
HMI tags "Consumtion"
   "DB_Zaehler_Anzeige_ViewPreShift" : Bool = PLC DB_Zaehler_Anzeige.ViewPreShift AT %DB211.DBX4.4, 1 s
   "DB_Zaehler_Anzeige_ReadWriteDeviceNo" : Int = PLC DB_Zaehler_Anzeige.ReadWriteDeviceNo AT %DB211.DBW0, 1 s
   "DB_Zaehler_Anzeige_Gesamt_Anzahl" : Int = PLC DB_Zaehler_Anzeige.Gesamt.Anzahl AT %DB211.DBW6, 1 s
   "DB_Zaehler_Anzeige_Gesamt_Verbrauch_K1" : Real = PLC DB_Zaehler_Anzeige.Gesamt.Verbrauch_K1 AT %DB211.DBD8, 1 s
   "DB_Zaehler_Anzeige_Gesamt_Verbrauch_K2" : Real = PLC DB_Zaehler_Anzeige.Gesamt.Verbrauch_K2 AT %DB211.DBD12, 1 s
   "DB_Zaehler_Anzeige_Gesamt_Verbrauch_K3" : Real = PLC DB_Zaehler_Anzeige.Gesamt.Verbrauch_K3 AT %DB211.DBD16, 1 s
   "DB_Zaehler_Anzeige_Gesamt_Verbrauch_K4" : Real = PLC DB_Zaehler_Anzeige.Gesamt.Verbrauch_K4 AT %DB211.DBD20, 1 s
   "DB_Zaehler_Anzeige_Gesamt_Verbrauch_K5" : Real = PLC DB_Zaehler_Anzeige.Gesamt.Verbrauch_K5 AT %DB211.DBD24, 1 s
   "DB_Zaehler_Anzeige_Gesamt_Verbrauch_K6" : Real = PLC DB_Zaehler_Anzeige.Gesamt.Verbrauch_K6 AT %DB211.DBD28, 1 s
   "DB_Zaehler_Anzeige_Gesamt_Verbrauch_K7" : Real = PLC DB_Zaehler_Anzeige.Gesamt.Verbrauch_K7 AT %DB211.DBD32, 1 s
   "DB_Zaehler_Anzeige_Gesamt_Verbrauch_K8" : Real = PLC DB_Zaehler_Anzeige.Gesamt.Verbrauch_K8 AT %DB211.DBD36, 1 s
   "DB_Zaehler_Anzeige_Counter{1}_Anzahl" : Int = PLC DB_Zaehler_Anzeige.Counter[1].Anzahl AT %DB211.DBW40, 1 s
   "DB_Zaehler_Anzeige_Counter{1}_Verbrauch_K1" : Real = PLC DB_Zaehler_Anzeige.Counter[1].Verbrauch_K1 AT %DB211.DBD42, 1 s
   "DB_Zaehler_Anzeige_Counter{1}_Verbrauch_K2" : Real = PLC DB_Zaehler_Anzeige.Counter[1].Verbrauch_K2 AT %DB211.DBD46, 1 s
   "DB_Zaehler_Anzeige_Counter{1}_Verbrauch_K3" : Real = PLC DB_Zaehler_Anzeige.Counter[1].Verbrauch_K3 AT %DB211.DBD50, 1 s
   "DB_Zaehler_Anzeige_Counter{1}_Verbrauch_K4" : Real = PLC DB_Zaehler_Anzeige.Counter[1].Verbrauch_K4 AT %DB211.DBD54, 1 s
   "DB_Zaehler_Anzeige_Counter{2}_Anzahl" : Int = PLC DB_Zaehler_Anzeige.Counter[2].Anzahl AT %DB211.DBW74, 1 s
   "DB_Zaehler_Anzeige_Counter{2}_Verbrauch_K1" : Real = PLC DB_Zaehler_Anzeige.Counter[2].Verbrauch_K1 AT %DB211.DBD76, 1 s
   "DB_Zaehler_Anzeige_Counter{2}_Verbrauch_K2" : Real = PLC DB_Zaehler_Anzeige.Counter[2].Verbrauch_K2 AT %DB211.DBD80, 1 s
   "DB_Zaehler_Anzeige_Counter{2}_Verbrauch_K3" : Real = PLC DB_Zaehler_Anzeige.Counter[2].Verbrauch_K3 AT %DB211.DBD84, 1 s
   "DB_Zaehler_Anzeige_Counter{2}_Verbrauch_K4" : Real = PLC DB_Zaehler_Anzeige.Counter[2].Verbrauch_K4 AT %DB211.DBD88, 1 s
   "DB_Zaehler_Anzeige_Counter{3}_Anzahl" : Int = PLC DB_Zaehler_Anzeige.Counter[3].Anzahl AT %DB211.DBW108, 1 s
   "DB_Zaehler_Anzeige_Counter{3}_Verbrauch_K1" : Real = PLC DB_Zaehler_Anzeige.Counter[3].Verbrauch_K1 AT %DB211.DBD110, 1 s
   "DB_Zaehler_Anzeige_Counter{3}_Verbrauch_K2" : Real = PLC DB_Zaehler_Anzeige.Counter[3].Verbrauch_K2 AT %DB211.DBD114, 1 s
   "DB_Zaehler_Anzeige_Counter{3}_Verbrauch_K3" : Real = PLC DB_Zaehler_Anzeige.Counter[3].Verbrauch_K3 AT %DB211.DBD118, 1 s
   "DB_Zaehler_Anzeige_Counter{3}_Verbrauch_K4" : Real = PLC DB_Zaehler_Anzeige.Counter[3].Verbrauch_K4 AT %DB211.DBD122, 1 s
   "DB_Zaehler_Anzeige_Counter{4}_Anzahl" : Int = PLC DB_Zaehler_Anzeige.Counter[4].Anzahl AT %DB211.DBW142, 1 s
   "DB_Zaehler_Anzeige_Counter{4}_Verbrauch_K1" : Real = PLC DB_Zaehler_Anzeige.Counter[4].Verbrauch_K1 AT %DB211.DBD144, 1 s
   "DB_Zaehler_Anzeige_Counter{4}_Verbrauch_K2" : Real = PLC DB_Zaehler_Anzeige.Counter[4].Verbrauch_K2 AT %DB211.DBD148, 1 s
   "DB_Zaehler_Anzeige_Counter{4}_Verbrauch_K3" : Real = PLC DB_Zaehler_Anzeige.Counter[4].Verbrauch_K3 AT %DB211.DBD152, 1 s
   "DB_Zaehler_Anzeige_Counter{4}_Verbrauch_K4" : Real = PLC DB_Zaehler_Anzeige.Counter[4].Verbrauch_K4 AT %DB211.DBD156, 1 s
   "DB_Zaehler_Anzeige_Counter{5}_Anzahl" : Int = PLC DB_Zaehler_Anzeige.Counter[5].Anzahl AT %DB211.DBW176, 1 s
   "DB_Zaehler_Anzeige_Counter{5}_Verbrauch_K1" : Real = PLC DB_Zaehler_Anzeige.Counter[5].Verbrauch_K1 AT %DB211.DBD178, 1 s
   "DB_Zaehler_Anzeige_Counter{5}_Verbrauch_K2" : Real = PLC DB_Zaehler_Anzeige.Counter[5].Verbrauch_K2 AT %DB211.DBD182, 1 s
   "DB_Zaehler_Anzeige_Counter{5}_Verbrauch_K3" : Real = PLC DB_Zaehler_Anzeige.Counter[5].Verbrauch_K3 AT %DB211.DBD186, 1 s
   "DB_Zaehler_Anzeige_Counter{5}_Verbrauch_K4" : Real = PLC DB_Zaehler_Anzeige.Counter[5].Verbrauch_K4 AT %DB211.DBD190, 1 s
   "DB_Zaehler_Anzeige_Counter{6}_Anzahl" : Int = PLC DB_Zaehler_Anzeige.Counter[6].Anzahl AT %DB211.DBW210, 1 s
   "DB_Zaehler_Anzeige_Counter{6}_Verbrauch_K1" : Real = PLC DB_Zaehler_Anzeige.Counter[6].Verbrauch_K1 AT %DB211.DBD212, 1 s
   "DB_Zaehler_Anzeige_Counter{6}_Verbrauch_K2" : Real = PLC DB_Zaehler_Anzeige.Counter[6].Verbrauch_K2 AT %DB211.DBD216, 1 s
   "DB_Zaehler_Anzeige_Counter{6}_Verbrauch_K3" : Real = PLC DB_Zaehler_Anzeige.Counter[6].Verbrauch_K3 AT %DB211.DBD220, 1 s
   "DB_Zaehler_Anzeige_Counter{6}_Verbrauch_K4" : Real = PLC DB_Zaehler_Anzeige.Counter[6].Verbrauch_K4 AT %DB211.DBD224, 1 s
   "DB_Zaehler_Anzeige_Counter{7}_Anzahl" : Int = PLC DB_Zaehler_Anzeige.Counter[7].Anzahl AT %DB211.DBW244, 1 s
   "DB_Zaehler_Anzeige_Counter{7}_Verbrauch_K1" : Real = PLC DB_Zaehler_Anzeige.Counter[7].Verbrauch_K1 AT %DB211.DBD246, 1 s
   "DB_Zaehler_Anzeige_Counter{7}_Verbrauch_K2" : Real = PLC DB_Zaehler_Anzeige.Counter[7].Verbrauch_K2 AT %DB211.DBD250, 1 s
   "DB_Zaehler_Anzeige_Counter{7}_Verbrauch_K3" : Real = PLC DB_Zaehler_Anzeige.Counter[7].Verbrauch_K3 AT %DB211.DBD254, 1 s
   "DB_Zaehler_Anzeige_Counter{7}_Verbrauch_K4" : Real = PLC DB_Zaehler_Anzeige.Counter[7].Verbrauch_K4 AT %DB211.DBD258, 1 s
   "DB_Zaehler_Anzeige_Counter{8}_Anzahl" : Int = PLC DB_Zaehler_Anzeige.Counter[8].Anzahl AT %DB211.DBW278, 1 s
   "DB_Zaehler_Anzeige_Counter{8}_Verbrauch_K1" : Real = PLC DB_Zaehler_Anzeige.Counter[8].Verbrauch_K1 AT %DB211.DBD280, 1 s
   "DB_Zaehler_Anzeige_Counter{8}_Verbrauch_K2" : Real = PLC DB_Zaehler_Anzeige.Counter[8].Verbrauch_K2 AT %DB211.DBD284, 1 s
   "DB_Zaehler_Anzeige_Counter{8}_Verbrauch_K3" : Real = PLC DB939_Tool_alloc_HMI.Alloc_stationTool[19] AT %DB211.DBD288, 1 s
   "DB_Zaehler_Anzeige_Counter{8}_Verbrauch_K4" : Real = PLC DB_Zaehler_Anzeige.Counter[8].Verbrauch_K4 AT %DB211.DBD292, 1 s
   "DB_Zaehler_Anzeige_Counter{9}_Anzahl" : Int = PLC DB_Zaehler_Anzeige.Counter[9].Anzahl AT %DB211.DBW312, 1 s
   "DB_Zaehler_Anzeige_Counter{9}_Verbrauch_K1" : Real = PLC DB_Zaehler_Anzeige.Counter[9].Verbrauch_K1 AT %DB211.DBD314, 1 s
   "DB_Zaehler_Anzeige_Counter{9}_Verbrauch_K2" : Real = PLC DB_Zaehler_Anzeige.Counter[9].Verbrauch_K2 AT %DB211.DBD318, 1 s
   "DB_Zaehler_Anzeige_Counter{9}_Verbrauch_K3" : Real = PLC DB_Zaehler_Anzeige.Counter[9].Verbrauch_K3 AT %DB211.DBD322, 1 s
   "DB_Zaehler_Anzeige_Counter{9}_Verbrauch_K4" : Real = PLC DB_Zaehler_Anzeige.Counter[9].Verbrauch_K4 AT %DB211.DBD326, 1 s
   "DB_Zaehler_Anzeige_Counter{10}_Anzahl" : Int = PLC DB_Zaehler_Anzeige.Counter[10].Anzahl AT %DB211.DBW346, 1 s
   "DB_Zaehler_Anzeige_Counter{10}_Verbrauch_K1" : Real = PLC DB_Zaehler_Anzeige.Counter[10].Verbrauch_K1 AT %DB211.DBD348, 1 s
   "DB_Zaehler_Anzeige_Counter{10}_Verbrauch_K2" : Real = PLC DB_Zaehler_Anzeige.Counter[10].Verbrauch_K2 AT %DB211.DBD352, 1 s
   "DB_Zaehler_Anzeige_Counter{10}_Verbrauch_K3" : Real = PLC DB_Zaehler_Anzeige.Counter[10].Verbrauch_K3 AT %DB211.DBD356, 1 s
   "DB_Zaehler_Anzeige_Counter{10}_Verbrauch_K4" : Real = PLC DB_Zaehler_Anzeige.Counter[10].Verbrauch_K4 AT %DB211.DBD360, 1 s
   "Consumtion_Name_1" : WString[10], internal
   "Consumtion_Name_2" : WString[10] AT %DB1.DBX0.0
   "Consumtion_Name_3" : WString[10] AT %DB1.DBX0.0
   "Consumtion_Name_4" : WString[10] AT %DB1.DBX0.0
   "Consumtion_Name_5" : WString[10] AT %DB1.DBX0.0
   "Consumtion_Name_6" : WString[10] AT %DB1.DBX0.0
   "Consumtion_Name_7" : WString[10] AT %DB1.DBX0.0
   "Consumtion_Name_8" : WString[10] AT %DB1.DBX0.0
   "Consumtion_Name_9" : WString[10] AT %DB1.DBX0.0
   "Consumtion_Name_10" : WString[10] AT %DB1.DBX0.0

HMI tags "Shift"
   "Shift1_Monday" : DateTime AT %DB1.DBX0.0
   "Shift1_Tuesday" : DateTime, internal
   "Shift1_Wenesday" : DateTime, internal
   "Shift1_Thrusday" : DateTime, internal
   "Shift1_Friday" : DateTime, internal
   "Shift1_Saturday" : DateTime, internal
   "Shift1_Sunday" : DateTime, internal
   "Shift2_Monday" : DateTime, internal
   "Shift2_Tuesday" : DateTime, internal
   "Shift2_Wenesday" : DateTime, internal
   "Shift2_Thrusday" : DateTime, internal
   "Shift2_Friday" : DateTime, internal
   "Shift2_Saturday" : DateTime, internal
   "Shift2_Sunday" : DateTime, internal
   "Shift3_Monday" : DateTime, internal
   "Shift3_Tuesday" : DateTime, internal
   "Shift3_Wenesday" : DateTime, internal
   "Shift3_Thrusday" : DateTime, internal
   "Shift3_Friday" : DateTime, internal
   "Shift3_Saturday" : DateTime, internal
   "Shift3_Sunday" : DateTime, internal
   "Shift4_Monday" : DateTime, internal
   "Shift4_Tuesday" : DateTime, internal
   "Shift4_Wenesday" : DateTime, internal
   "Shift4_Thrusday" : DateTime, internal
   "Shift4_Friday" : DateTime, internal
   "Shift4_Saturday" : DateTime, internal
   "Shift4_Sunday" : DateTime, internal
   "Check_Shift1_Monday" : Bool, internal
   "Check_Shift1_Tuesday" : Bool, internal
   "Check_Shift1_Wenesday" : Bool, internal
   "Check_Shift1_Thrusday" : Bool, internal
   "Check_Shift1_Friday" : Bool, internal
   "Check_Shift1_Saturday" : Bool, internal
   "Check_Shift1_Sunday" : Bool, internal
   "Check_Shift2_Monday" : Bool, internal
   "Check_Shift2_Tuesday" : Bool, internal
   "Check_Shift2_Wenesday" : Bool, internal
   "Check_Shift2_Thrusday" : Bool, internal
   "Check_Shift2_Friday" : Bool, internal
   "Check_Shift2_Saturday" : Bool, internal
   "Check_Shift2_Sunday" : Bool, internal
   "Check_Shift3_Monday" : Bool, internal
   "Check_Shift3_Tuesday" : Bool, internal
   "Check_Shift3_Wenesday" : Bool, internal
   "Check_Shift3_Thrusday" : Bool, internal
   "Check_Shift3_Friday" : Bool, internal
   "Check_Shift3_Saturday" : Bool, internal
   "Check_Shift3_Sunday" : Bool, internal
   "Check_Shift4_Monday" : Bool, internal
   "Check_Shift4_Tuesday" : Bool, internal
   "Check_Shift4_Wenesday" : Bool, internal
   "Check_Shift4_Thrusday" : Bool, internal
   "Check_Shift4_Friday" : Bool, internal
   "Check_Shift4_Saturday" : Bool, internal
   "Check_Shift4_Sunday" : Bool, internal
   "Shift_Protocol_1" : DateTime, internal
      on ChangeValue: function_f38ba6b2("ShiftProtocol", U 1, 1, 0, N)
   "Shift_Protocol_2" : DateTime, internal
      on ChangeValue: function_f38ba6b2("ShiftProtocol", U 1, 1, 0, N)
   "Shift_Protocol_3" : DateTime, internal
      on ChangeValue: function_f38ba6b2("ShiftProtocol", U 1, 1, 0, N)
   "Shift_Protocol_4" : DateTime, internal
      on ChangeValue: function_f38ba6b2("ShiftProtocol", U 1, 1, 0, N)
   "Shift_Protocol_5" : DateTime, internal
      on ChangeValue: function_f38ba6b2("ShiftProtocol", U 1, 1, 0, N)
   "Shift_Protocol_6" : DateTime, internal
      on ChangeValue: function_f38ba6b2("ShiftProtocol", U 1, 1, 0, N)
   "Shift_Protocol_7" : DateTime, internal
      on ChangeValue: function_f38ba6b2("ShiftProtocol", U 1, 1, 0, N)
   "Shift_Protocol_8" : DateTime, internal
      on ChangeValue: function_f38ba6b2("ShiftProtocol", U 1, 1, 0, N)
   "Shift_Protocol_9" : DateTime, internal
      on ChangeValue: function_f38ba6b2("ShiftProtocol", U 1, 1, 0, N)
   "Shift_Protocol_10" : DateTime, internal
      on ChangeValue: function_f38ba6b2("ShiftProtocol", U 1, 1, 0, N)
   "Shift_Protocol_11" : DateTime, internal
      on ChangeValue: function_f38ba6b2("ShiftProtocol", U 1, 1, 0, N)
   "Shift_Protocol_12" : DateTime, internal
      on ChangeValue: function_f38ba6b2("ShiftProtocol", U 1, 1, 0, N)
   "Shift_Protocol_13" : DateTime, internal
      on ChangeValue: function_f38ba6b2("ShiftProtocol", U 1, 1, 0, N)
   "Shift_Protocol_14" : DateTime, internal
      on ChangeValue: function_f38ba6b2("ShiftProtocol", U 1, 1, 0, N)
   "Shift_Protocol_15" : DateTime, internal
      on ChangeValue: function_f38ba6b2("ShiftProtocol", U 1, 1, 0, N)
   "Shift_Protocol_16" : DateTime, internal
      on ChangeValue: function_f38ba6b2("ShiftProtocol", U 1, 1, 0, N)
   "Shift_Protocol_17" : DateTime, internal
      on ChangeValue: function_f38ba6b2("ShiftProtocol", U 1, 1, 0, N)
   "Shift_Protocol_18" : DateTime, internal
      on ChangeValue: function_f38ba6b2("ShiftProtocol", U 1, 1, 0, N)
   "Shift_Protocol_19" : DateTime, internal
      on ChangeValue: function_f38ba6b2("ShiftProtocol", U 1, 1, 0, N)
   "Shift_Protocol_20" : DateTime, internal
      on ChangeValue: function_f38ba6b2("ShiftProtocol", U 1, 1, 0, N)
   "Shift_Protocol_21" : DateTime, internal
      on ChangeValue: function_f38ba6b2("ShiftProtocol", U 1, 1, 0, N)
   "Next shift" : DateTime, internal
   "Shift_1_1" : DateTime, internal
   "Shift_1_2" : DateTime, internal
   "Shift_1_3" : DateTime, internal
   "Shift_1_4" : DateTime, internal
   "Shift_2_1" : DateTime, internal
   "Shift_2_2" : DateTime, internal
   "Shift_2_3" : DateTime, internal
   "Shift_2_4" : DateTime, internal
   "Shift_3_1" : DateTime, internal
   "Shift_3_2" : DateTime, internal
   "Shift_3_3" : DateTime, internal
   "Shift_3_4" : DateTime, internal
   "Shift_4_1" : DateTime, internal
   "Shift_4_2" : DateTime, internal
   "Shift_4_3" : DateTime, internal
   "Shift_4_4" : DateTime, internal
   "Shift_5_1" : DateTime, internal
   "Shift_5_2" : DateTime, internal
   "Shift_5_3" : DateTime, internal
   "Shift_5_4" : DateTime, internal
   "Shift_6_1" : DateTime, internal
   "Shift_6_2" : DateTime, internal
   "Shift_6_3" : DateTime, internal
   "Shift_6_4" : DateTime, internal
   "Shift_7_1" : DateTime, internal
   "Shift_7_2" : DateTime, internal
   "Shift_7_3" : DateTime, internal
   "Shift_7_4" : DateTime, internal
   "Shift_En_1_1" : Bool, internal
   "Shift_En_1_2" : Bool, internal
   "Shift_En_1_3" : Bool, internal
   "Shift_En_1_4" : Bool, internal
   "Shift_En_2_1" : Bool, internal
   "Shift_En_2_2" : Bool, internal
   "Shift_En_2_3" : Bool, internal
   "Shift_En_2_4" : Bool, internal
   "Shift_En_3_1" : Bool, internal
   "Shift_En_3_2" : Bool, internal
   "Shift_En_3_3" : Bool, internal
   "Shift_En_3_4" : Bool, internal
   "Shift_En_4_1" : Bool, internal
   "Shift_En_4_2" : Bool, internal
   "Shift_En_4_3" : Bool, internal
   "Shift_En_4_4" : Bool, internal
   "Shift_En_5_1" : Bool, internal
   "Shift_En_5_2" : Bool, internal
   "Shift_En_5_3" : Bool, internal
   "Shift_En_5_4" : Bool, internal
   "Shift_En_6_1" : Bool, internal
   "Shift_En_6_2" : Bool, internal
   "Shift_En_6_3" : Bool, internal
   "Shift_En_6_4" : Bool, internal
   "Shift_En_7_1" : Bool, internal
   "Shift_En_7_2" : Bool, internal
   "Shift_En_7_3" : Bool, internal
   "Shift_En_7_4" : Bool, internal

HMI tags "ToolAllocation"
   "DB939_Tool_alloc_HMI_Alloc_stationTool{1}" : Int = PLC DB939_Tool_alloc_HMI.Alloc_stationTool[1], 1 s
   "DB939_Tool_alloc_HMI_Alloc_stationTool{2}" : Int = PLC DB939_Tool_alloc_HMI.Alloc_stationTool[2], 1 s
   "DB939_Tool_alloc_HMI_Alloc_stationTool{3}" : Int = PLC DB939_Tool_alloc_HMI.Alloc_stationTool[3], 1 s
   "DB939_Tool_alloc_HMI_Alloc_stationTool{4}" : Int = PLC DB939_Tool_alloc_HMI.Alloc_stationTool[4], 1 s
   "DB939_Tool_alloc_HMI_Alloc_stationTool{5}" : Int = PLC DB939_Tool_alloc_HMI.Alloc_stationTool[5], 1 s
   "DB939_Tool_alloc_HMI_Alloc_stationTool{6}" : Int = PLC DB939_Tool_alloc_HMI.Alloc_stationTool[6], 1 s
   "DB939_Tool_alloc_HMI_Alloc_stationTool{7}" : Int = PLC DB939_Tool_alloc_HMI.Alloc_stationTool[7], 1 s
   "DB939_Tool_alloc_HMI_Alloc_stationTool{8}" : Int = PLC DB939_Tool_alloc_HMI.Alloc_stationTool[8], 1 s
   "DB939_Tool_alloc_HMI_Alloc_stationTool{9}" : Int = PLC DB939_Tool_alloc_HMI.Alloc_stationTool[9], 1 s
   "DB939_Tool_alloc_HMI_Alloc_stationTool{10}" : Int = PLC DB939_Tool_alloc_HMI.Alloc_stationTool[10], 1 s
   "DB939_Tool_alloc_HMI_Alloc_stationTool{11}" : Int = PLC DB939_Tool_alloc_HMI.Alloc_stationTool[11], 1 s
   "DB939_Tool_alloc_HMI_Alloc_stationTool{12}" : Int = PLC DB939_Tool_alloc_HMI.Alloc_stationTool[12], 1 s
   "DB939_Tool_alloc_HMI_Alloc_stationTool{13}" : Int = PLC DB939_Tool_alloc_HMI.Alloc_stationTool[13], 1 s
   "DB939_Tool_alloc_HMI_Alloc_stationTool{14}" : Int = PLC DB939_Tool_alloc_HMI.Alloc_stationTool[14], 1 s
   "DB939_Tool_alloc_HMI_Alloc_stationTool{15}" : Int = PLC DB939_Tool_alloc_HMI.Alloc_stationTool[15], 1 s
   "DB939_Tool_alloc_HMI_Alloc_stationTool{16}" : Int = PLC DB939_Tool_alloc_HMI.Alloc_stationTool[16], 1 s
   "DB939_Tool_alloc_HMI_Alloc_stationTool{17}" : Int = PLC DB939_Tool_alloc_HMI.Alloc_stationTool[17], 1 s
   "DB939_Tool_alloc_HMI_Alloc_stationTool{18}" : Int = PLC DB939_Tool_alloc_HMI.Alloc_stationTool[18], 1 s
   "DB939_Tool_alloc_HMI_Alloc_stationTool{19}" : Int = PLC DB939_Tool_alloc_HMI.Alloc_stationTool[19], 1 s
   "DB939_Tool_alloc_HMI_Alloc_stationTool{20}" : Int = PLC DB939_Tool_alloc_HMI.Alloc_stationTool[20], 1 s
   "DB939_Tool_alloc_HMI_Alloc_stationTool{21}" : Int = PLC DB939_Tool_alloc_HMI.Alloc_stationTool[21], 1 s
   "DB939_Tool_alloc_HMI_Alloc_stationTool{22}" : Int = PLC DB939_Tool_alloc_HMI.Alloc_stationTool[22], 1 s
   "DB939_Tool_alloc_HMI_Alloc_stationTool{23}" : Int = PLC DB939_Tool_alloc_HMI.Alloc_stationTool[23], 1 s
   "DB939_Tool_alloc_HMI_Alloc_stationTool{24}" : Int = PLC DB939_Tool_alloc_HMI.Alloc_stationTool[24], 1 s
   "DB939_Tool_alloc_HMI_Alloc_stationTool{25}" : Int = PLC DB939_Tool_alloc_HMI.Alloc_stationTool[25], 1 s
   "DB939_Tool_alloc_HMI_Alloc_stationTool{26}" : Int = PLC DB939_Tool_alloc_HMI.Alloc_stationTool[26], 1 s
   "DB939_Tool_alloc_HMI_Alloc_stationTool{27}" : Int = PLC DB939_Tool_alloc_HMI.Alloc_stationTool[27], 1 s
   "DB939_Tool_alloc_HMI_Alloc_stationTool{28}" : Int = PLC DB939_Tool_alloc_HMI.Alloc_stationTool[28], 1 s
   "DB939_Tool_alloc_HMI_Alloc_stationTool{29}" : Int = PLC DB939_Tool_alloc_HMI.Alloc_stationTool[29], 1 s
   "DB939_Tool_alloc_HMI_Alloc_stationTool{30}" : Int = PLC DB939_Tool_alloc_HMI.Alloc_stationTool[30], 1 s
   "DB939_Tool_alloc_HMI_Alloc_tool_name{1}" : String[20] = PLC DB939_Tool_alloc_HMI.Alloc_tool_name[1], 1 s
   "DB939_Tool_alloc_HMI_Alloc_tool_name{2}" : String[20] = PLC DB939_Tool_alloc_HMI.Alloc_tool_name[2], 1 s
   "DB939_Tool_alloc_HMI_Alloc_tool_name{3}" : String[20] = PLC DB939_Tool_alloc_HMI.Alloc_tool_name[3], 1 s
   "DB939_Tool_alloc_HMI_Alloc_tool_name{4}" : String[20] = PLC DB939_Tool_alloc_HMI.Alloc_tool_name[4], 1 s
   "DB939_Tool_alloc_HMI_Alloc_tool_name{5}" : String[20] = PLC DB939_Tool_alloc_HMI.Alloc_tool_name[5], 1 s
   "DB939_Tool_alloc_HMI_Alloc_tool_name{6}" : String[20] = PLC DB939_Tool_alloc_HMI.Alloc_tool_name[6], 1 s
   "DB939_Tool_alloc_HMI_Alloc_tool_name{7}" : String[20] = PLC DB939_Tool_alloc_HMI.Alloc_tool_name[7], 1 s
   "DB939_Tool_alloc_HMI_Alloc_tool_name{8}" : String[20] = PLC DB939_Tool_alloc_HMI.Alloc_tool_name[8], 1 s
   "DB939_Tool_alloc_HMI_Alloc_tool_name{9}" : String[20] = PLC DB939_Tool_alloc_HMI.Alloc_tool_name[9], 1 s
   "DB939_Tool_alloc_HMI_Alloc_tool_name{10}" : String[20] = PLC DB939_Tool_alloc_HMI.Alloc_tool_name[10], 1 s
   "DB939_Tool_alloc_HMI_Alloc_tool_name{11}" : String[20] = PLC DB939_Tool_alloc_HMI.Alloc_tool_name[11], 1 s
   "DB939_Tool_alloc_HMI_Alloc_tool_name{12}" : String[20] = PLC DB939_Tool_alloc_HMI.Alloc_tool_name[12], 1 s
   "DB939_Tool_alloc_HMI_Alloc_tool_name{13}" : String[20] = PLC DB939_Tool_alloc_HMI.Alloc_tool_name[13], 1 s
   "DB939_Tool_alloc_HMI_Alloc_tool_name{14}" : String[20] = PLC DB939_Tool_alloc_HMI.Alloc_tool_name[14], 1 s
   "DB939_Tool_alloc_HMI_Alloc_tool_name{15}" : String[20] = PLC DB939_Tool_alloc_HMI.Alloc_tool_name[15], 1 s
   "DB939_Tool_alloc_HMI_Alloc_tool_name{16}" : String[20] = PLC DB939_Tool_alloc_HMI.Alloc_tool_name[16], 1 s
   "DB939_Tool_alloc_HMI_Alloc_tool_name{17}" : String[20] = PLC DB939_Tool_alloc_HMI.Alloc_tool_name[17], 1 s
   "DB939_Tool_alloc_HMI_Alloc_tool_name{18}" : String[20] = PLC DB939_Tool_alloc_HMI.Alloc_tool_name[18], 1 s
   "DB939_Tool_alloc_HMI_Alloc_tool_name{19}" : String[20] = PLC DB939_Tool_alloc_HMI.Alloc_tool_name[19], 1 s
   "DB939_Tool_alloc_HMI_Alloc_tool_name{20}" : String[20] = PLC DB939_Tool_alloc_HMI.Alloc_tool_name[20], 1 s
   "DB939_Tool_alloc_HMI_Alloc_tool_name{21}" : String[20] = PLC DB939_Tool_alloc_HMI.Alloc_tool_name[21], 1 s
   "DB939_Tool_alloc_HMI_Alloc_tool_name{22}" : String[20] = PLC DB939_Tool_alloc_HMI.Alloc_tool_name[22], 1 s
   "DB939_Tool_alloc_HMI_Alloc_tool_name{23}" : String[20] = PLC DB939_Tool_alloc_HMI.Alloc_tool_name[23], 1 s
   "DB939_Tool_alloc_HMI_Alloc_tool_name{24}" : String[20] = PLC DB939_Tool_alloc_HMI.Alloc_tool_name[24], 1 s
   "DB939_Tool_alloc_HMI_Alloc_tool_name{25}" : String[20] = PLC DB939_Tool_alloc_HMI.Alloc_tool_name[25], 1 s
   "DB939_Tool_alloc_HMI_Alloc_tool_name{26}" : String[20] = PLC DB939_Tool_alloc_HMI.Alloc_tool_name[26], 1 s
   "DB939_Tool_alloc_HMI_Alloc_tool_name{27}" : String[20] = PLC DB939_Tool_alloc_HMI.Alloc_tool_name[27], 1 s
   "DB939_Tool_alloc_HMI_Alloc_tool_name{28}" : String[20] = PLC DB939_Tool_alloc_HMI.Alloc_tool_name[28], 1 s
   "DB939_Tool_alloc_HMI_Alloc_tool_name{29}" : String[20] = PLC DB939_Tool_alloc_HMI.Alloc_tool_name[29], 1 s
   "DB939_Tool_alloc_HMI_Alloc_tool_name{30}" : String[20] = PLC DB939_Tool_alloc_HMI.Alloc_tool_name[30], 1 s
   "DB939_Tool_alloc_HMI_AllocList_page" : Int = PLC DB939_Tool_alloc_HMI.AllocList_page AT %DB1.DBX0.0, 1 s
   "DB939_Tool_alloc_HMI_Selected_prog" : Int = PLC DB939_Tool_alloc_HMI.Selected_prog AT %DB1.DBX0.0, 1 s
   "DB939_Tool_alloc_HMI_Select_hand_automatic_alloc" : Bool = PLC DB939_Tool_alloc_HMI.Select_hand_automatic_alloc, 1 s
   "DB939_Tool_alloc_HMI_MH_No_selected" : Int = PLC DB939_Tool_alloc_HMI.MH_No_selected, 1 s
      on ChangeValue: "ToolAllocation_Sec"()
      on AboveUpperLimit: "ToolAllocation_Sec"()
   "DB939_Tool_alloc_HMI_Limit_allocation_list" : Int = PLC DB939_Tool_alloc_HMI.Limit_allocation_list, 1 s
   "DB939_Tool_alloc_HMI_SaveSortProgs{1}" : Int = PLC DB939_Tool_alloc_HMI.SaveSortProgs[1], 1 s
   "DB939_Tool_alloc_HMI_SaveSortProgs{2}" : Int = PLC DB939_Tool_alloc_HMI.SaveSortProgs[2], 1 s
   "DB939_Tool_alloc_HMI_SaveSortProgs{3}" : Int = PLC DB939_Tool_alloc_HMI.SaveSortProgs[3], 1 s
   "DB939_Tool_alloc_HMI_SaveSortProgs{4}" : Int = PLC DB939_Tool_alloc_HMI.SaveSortProgs[4], 1 s
   "DB939_Tool_alloc_HMI_SaveSortProgs{5}" : Int = PLC DB939_Tool_alloc_HMI.SaveSortProgs[5], 1 s
   "DB939_Tool_alloc_HMI_SaveSortProgs{6}" : Int = PLC DB939_Tool_alloc_HMI.SaveSortProgs[6], 1 s
   "DB939_Tool_alloc_HMI_SaveSortProgs{7}" : Int = PLC DB939_Tool_alloc_HMI.SaveSortProgs[7], 1 s
   "DB939_Tool_alloc_HMI_SaveSortProgs{8}" : Int = PLC DB939_Tool_alloc_HMI.SaveSortProgs[8], 1 s
   "DB939_Tool_alloc_HMI_SaveSortProgs{9}" : Int = PLC DB939_Tool_alloc_HMI.SaveSortProgs[9], 1 s
   "DB939_Tool_alloc_HMI_SaveSortProgs{10}" : Int = PLC DB939_Tool_alloc_HMI.SaveSortProgs[10], 1 s
   "DB939_Tool_alloc_HMI_SaveSortProgs{11}" : Int = PLC DB939_Tool_alloc_HMI.SaveSortProgs[11], 1 s
   "DB939_Tool_alloc_HMI_SaveSortProgs{12}" : Int = PLC DB939_Tool_alloc_HMI.SaveSortProgs[12], 1 s
   "DB939_Tool_alloc_HMI_SaveSortProgs{13}" : Int = PLC DB939_Tool_alloc_HMI.SaveSortProgs[13], 1 s
   "DB939_Tool_alloc_HMI_SaveSortProgs{14}" : Int = PLC DB939_Tool_alloc_HMI.SaveSortProgs[14], 1 s
   "DB939_Tool_alloc_HMI_SaveSortProgs{15}" : Int = PLC DB939_Tool_alloc_HMI.SaveSortProgs[15], 1 s
   "DB939_Tool_alloc_HMI_SaveSortProgs{16}" : Int = PLC DB939_Tool_alloc_HMI.SaveSortProgs[16], 1 s
   "DB939_Tool_alloc_HMI_SaveSortProgs{17}" : Int = PLC DB939_Tool_alloc_HMI.SaveSortProgs[17], 1 s
   "DB939_Tool_alloc_HMI_SaveSortProgs{18}" : Int = PLC DB939_Tool_alloc_HMI.SaveSortProgs[18], 1 s
   "DB939_Tool_alloc_HMI_SaveSortProgs{19}" : Int = PLC DB939_Tool_alloc_HMI.SaveSortProgs[19], 1 s
   "DB939_Tool_alloc_HMI_SaveSortProgs{20}" : Int = PLC DB939_Tool_alloc_HMI.SaveSortProgs[20], 1 s
   "DB939_Tool_alloc_HMI_SaveSortProg_name{1}" : String[20] = PLC DB939_Tool_alloc_HMI.SaveSortProg_name[1], 1 s
   "DB939_Tool_alloc_HMI_SaveSortProg_name{2}" : String[20] = PLC DB939_Tool_alloc_HMI.SaveSortProg_name[2], 1 s
   "DB939_Tool_alloc_HMI_SaveSortProg_name{3}" : String[20] = PLC DB939_Tool_alloc_HMI.SaveSortProg_name[3], 1 s
   "DB939_Tool_alloc_HMI_SaveSortProg_name{4}" : String[20] = PLC DB939_Tool_alloc_HMI.SaveSortProg_name[4], 1 s
   "DB939_Tool_alloc_HMI_SaveSortProg_name{5}" : String[20] = PLC DB939_Tool_alloc_HMI.SaveSortProg_name[5], 1 s
   "DB939_Tool_alloc_HMI_SaveSortProg_name{6}" : String[20] = PLC DB939_Tool_alloc_HMI.SaveSortProg_name[6], 1 s
   "DB939_Tool_alloc_HMI_SaveSortProg_name{7}" : String[20] = PLC DB939_Tool_alloc_HMI.SaveSortProg_name[7], 1 s
   "DB939_Tool_alloc_HMI_SaveSortProg_name{8}" : String[20] = PLC DB939_Tool_alloc_HMI.SaveSortProg_name[8], 1 s
   "DB939_Tool_alloc_HMI_SaveSortProg_name{9}" : String[20] = PLC DB939_Tool_alloc_HMI.SaveSortProg_name[9], 1 s
   "DB939_Tool_alloc_HMI_SaveSortProg_name{10}" : String[20] = PLC DB939_Tool_alloc_HMI.SaveSortProg_name[10], 1 s
   "DB939_Tool_alloc_HMI_SaveSortProg_name{11}" : String[20] = PLC DB939_Tool_alloc_HMI.SaveSortProg_name[11], 1 s
   "DB939_Tool_alloc_HMI_SaveSortProg_name{12}" : String[20] = PLC DB939_Tool_alloc_HMI.SaveSortProg_name[12], 1 s
   "DB939_Tool_alloc_HMI_SaveSortProg_name{13}" : String[20] = PLC DB939_Tool_alloc_HMI.SaveSortProg_name[13], 1 s
   "DB939_Tool_alloc_HMI_SaveSortProg_name{14}" : String[20] = PLC DB939_Tool_alloc_HMI.SaveSortProg_name[14], 1 s
   "DB939_Tool_alloc_HMI_SaveSortProg_name{15}" : String[20] = PLC DB939_Tool_alloc_HMI.SaveSortProg_name[15], 1 s
   "DB939_Tool_alloc_HMI_SaveSortProg_name{16}" : String[20] = PLC DB939_Tool_alloc_HMI.SaveSortProg_name[16], 1 s
   "DB939_Tool_alloc_HMI_SaveSortProg_name{17}" : String[20] = PLC DB939_Tool_alloc_HMI.SaveSortProg_name[17], 1 s
   "DB939_Tool_alloc_HMI_SaveSortProg_name{18}" : String[20] = PLC DB939_Tool_alloc_HMI.SaveSortProg_name[18], 1 s
   "DB939_Tool_alloc_HMI_SaveSortProg_name{19}" : String[20] = PLC DB939_Tool_alloc_HMI.SaveSortProg_name[19], 1 s
   "DB939_Tool_alloc_HMI_SaveSortProg_name{20}" : String[20] = PLC DB939_Tool_alloc_HMI.SaveSortProg_name[20], 1 s
   "DB939_Tool_alloc_HMI_SavedProgs_decrease" : Bool = PLC DB939_Tool_alloc_HMI.SavedProgs_decrease AT %DB1.DBX0.0, 1 s
   "DB939_Tool_alloc_HMI_SavedProgs_increase" : Bool = PLC DB939_Tool_alloc_HMI.SavedProgs_increase AT %DB1.DBX0.0, 1 s
   "Tag_1" : Int = PLC DB939_Tool_alloc_HMI.Selected_SavedProg AT %DB1.DBX0.0, 1 s
   "DB939_Tool_alloc_HMI_Delete_selected_tool" : Int = PLC DB939_Tool_alloc_HMI.Delete_selected_tool, 1 s
   "DB939_Tool_alloc_HMI_SavedProgs_decrease_visible" : Bool = PLC DB939_Tool_alloc_HMI.SavedProgs_decrease_visible, 1 s
   "DB939_Tool_alloc_HMI_SavedProgs_increase_visible" : Bool = PLC DB939_Tool_alloc_HMI.SavedProgs_increase_visible, 1 s
   "DB939_Tool_alloc_HMI_Delete_tool_in _all_allocations" : Bool = PLC DB939_Tool_alloc_HMI."Delete_tool_in _all_allocations", 1 s

HMI tags "Internal_animation"
   "Tool_Allocation_Numb_1" : Int, internal
   "Tool_Allocation_Numb_2" : Int, internal
   "Tool_Allocation_Numb_3" : Int, internal
   "Tool_Allocation_Numb_4" : Int, internal
   "Tool_Allocation_Numb_5" : Int, internal
   "Tool_Allocation_Numb_6" : Int, internal
   "Tool_Allocation_Numb_7" : Int, internal
   "Tool_Allocation_Numb_8" : Int, internal
   "Tool_Allocation_Numb_9" : Int, internal
   "Tool_Allocation_Numb_10" : Int, internal
   "Tool_Allocation_Numb_11" : Int, internal
   "Tool_Allocation_Numb_12" : Int, internal
   "Tool_Allocation_Numb_13" : Int, internal
   "Tool_Allocation_Numb_14" : Int, internal
   "Tool_Allocation_Numb_15" : Int, internal
   "Tool_Allocation_Numb_16" : Int, internal
   "Tool_Allocation_Numb_17" : Int, internal
   "Tool_Allocation_Numb_18" : Int, internal
   "Tool_Allocation_Numb_19" : Int, internal
   "Tool_Allocation_Numb_20" : Int, internal
   "Tool_Allocation_Numb_21" : Int, internal
   "Tool_Allocation_Numb_22" : Int, internal
   "Tool_Allocation_Numb_23" : Int, internal
   "Tool_Allocation_Numb_24" : Int, internal
   "Tool_Allocation_Numb_25" : Int, internal
   "Tool_Allocation_Numb_26" : Int, internal
   "Tool_Allocation_Numb_27" : Int, internal
   "Tool_Allocation_Numb_28" : Int, internal
   "Tool_Allocation_Numb_29" : Int, internal
   "Tool_Allocation_Numb_30" : Int, internal
   "Tank_Visibility Control" : Int, internal
   "Recipe_Appearance_Control" : Int, internal
   "Consumtion_Numb_1" : Int, internal
   "Consumtion_Numb_2" : Int, internal
   "Consumtion_Numb_3" : Int, internal
   "Consumtion_Numb_4" : Int, internal
   "Consumtion_Numb_5" : Int, internal
   "Consumtion_Numb_6" : Int, internal
   "Consumtion_Numb_7" : Int, internal
   "Consumtion_Numb_8" : Int, internal
   "Consumtion_Numb_9" : Int, internal
   "Consumtion_Numb_10" : Int, internal
   "Part_Counter_Numb_1" : Int, internal
   "Part_Counter_Numb_2" : Int, internal
   "Part_Counter_Numb_3" : Int, internal
   "Part_Counter_Numb_4" : Int, internal
   "Part_Counter_Numb_5" : Int, internal
   "Part_Counter_Numb_6" : Int, internal
   "Part_Counter_Numb_7" : Int, internal
   "Part_Counter_Numb_8" : Int, internal
   "Part_Counter_Numb_9" : Int, internal
   "Part_Counter_Numb_10" : Int, internal
   "Part_Counter_Numb_11" : Int, internal
   "Part_Counter_Numb_12" : Int, internal
   "Part_Counter_Numb_13" : Int, internal
   "Part_Counter_Numb_14" : Int, internal
   "Part_Counter_Numb_15" : Int, internal
   "Part_Counter_Numb_16" : Int, internal
   "Part_Counter_Numb_17" : Int, internal
   "Part_Counter_Numb_18" : Int, internal
   "Part_Counter_Numb_19" : Int, internal
   "Part_Counter_Numb_20" : Int, internal
   "Part_Counter_Numb_21" : Int, internal
   "Part_Counter_Numb_22" : Int, internal
   "Part_Counter_Numb_23" : Int, internal
   "Part_Counter_Numb_24" : Int, internal
   "Part_Counter_Numb_25" : Int, internal
   "Part_Counter_Numb_26" : Int, internal
   "Part_Counter_Numb_27" : Int, internal
   "Part_Counter_Numb_28" : Int, internal
   "Part_Counter_Numb_29" : Int, internal
   "Part_Counter_Numb_30" : Int, internal
   "Create Part Counter Control" : Int, internal
   "Create Part Counter Button Save" : Int, internal
   "Create Part Counter Multiplexing Control" : Int, internal
   "Consumtion Name Multiplexing Control" : Int, internal
   "LargeScalleValues Control" : Int, internal
   "Archived Alarm Control" : Int, internal
   "First_Runtime_Rising_Control" : Int, internal
   "Internal_Tank_" : Int, internal
   "System Setting Screen Control" : Int, internal
   "OpenFileBrowserPath" : WString[30], internal
   "OpenFileBrowser_Status" : Int, internal
   "Robot Screen Visibility Control" : Int, internal
   "Logging_Visibility" : Int, internal
   "ImportDataFrom_SD" : WString[45], internal
   "ImportDataFrom_SD_stat" : Int, internal
   "Service Screen Control Visibility" : Int, internal
   "refresh_Alarm" : Int, internal
   "ImportDataFrom_USB_stat" : Int, internal
   "ImportDataFrom_USB" : WString[100], internal
   "R_date" : DateTime, internal
   "R_Time" : DateTime, internal
   "Archive Alarm Number" : Int, internal
   "Shift Protocol Alarm view_1" : Int, internal
   "Shift Protocol Alarm view_2" : Int, internal
   "Shift Protocol Alarm view_3" : Int, internal
   "Shift Protocol Alarm view_4" : Int, internal
   "Shift Protocol Alarm view_5" : Int, internal
   "Shift Protocol Alarm view_6" : Int, internal
   "Shift Protocol Alarm view_7" : Int, internal
   "Shift Protocol Alarm view_8" : Int, internal
   "Shift Protocol Alarm view_9" : Int, internal
   "Shift Protocol Alarm view_10" : Int, internal
   "Shift Protocol Alarm view_11" : Int, internal
   "Shift Protocol Alarm view_12" : Int, internal
   "Shift Protocol Alarm view_13" : Int, internal
   "Shift Protocol Alarm view_14" : Int, internal
   "Shift Protocol Alarm view_15" : Int, internal
   "Shift Protocol Alarm view_16" : Int, internal
   "Shift Protocol Alarm view_17" : Int, internal
   "Shift Protocol Alarm view_18" : Int, internal
   "Shift Protocol Alarm view_19" : Int, internal
   "Shift Protocol Alarm view_20" : Int, internal
   "Shift Protocol Alarm view_21" : Int, internal
   "CopyLogControl" : Int, internal
   "HMI_Tag_1(2)" : Bool, internal
   "ServiceScreenControl" : Int, internal
   "Nav_1" : Int, internal
   "Nav_2" : Int, internal
   "Nav_3" : Int, internal
   "Nav_4" : Int, internal
   "Nav_5" : Int, internal
   "Nav_6" : Int, internal
   "Nav_7" : Int, internal

